(* Logix 5000 project; controller FV vendor 1 type 14 code 217 rev 31.11; software revision 31.00; part 34 of 63 *)
(* tags used below, declared in another part *)
   CheckTimeMask : INT;
   CWD : CHECKWORD_FLAGS;
   Dummy : BOOL;
   FV_A_CTNo : DINT;
   FV_A_CTNo_PLCtoPC : DINT;
   FV_A_FVNo : DINT;
   FV_A_FVNo_PLCtoPC : DINT;
   FV_A_MVNo : DINT;
   FV_A_MVNo_PLCtoPC : DINT;
   FV_ALARM_RETURNED_STRING : STRING;
   FV_Event_Alarm_Tag : ALARM_DIGITAL;
   FV_Event_control_FIFO : CONTROL;
   FV_Event_control_FIFO_Operation_Type : CONTROL;
   FV_Event_Delay_For_Data : TIMER;
   FV_Event_Delay_For_PLC_Startup_Data : TIMER;
   FV_Event_Delay_Timer : TIMER;
   FV_Event_Delay_Timer_Off : TIMER;
   FV_Event_from_buffer : STRING;
   FV_Event_from_buffer_LogData1 : REAL;
   FV_Event_from_buffer_LogData2 : REAL;
   FV_Event_from_buffer_LogData3 : REAL;
   FV_Event_from_buffer_LogData4 : REAL;
   FV_Event_from_buffer_Operation_Type : DINT;
   fv_event_step : DINT;   // 0 - Wait For Event 1 - Sending Event To FactoryTalk 2 - Waiting For Delay Before Next Event Allowed
   FV_Event_String_Last : STRING;
   FV_Event_Transact_Trigger_Tag : DINT;
   FV_Events_FIFO_Buffer : STRING[31];
   FV_Events_FIFO_Buffer_Operation_Type : DINT[31];
   FV_Last_LogData_For_Op : REAL[30,20];
   FV_N20 : INT[255];   // YSVFILL<PC YSV Filling data fro m PC
   FV_N21 : INT[255];   // YSVFILL>PC YSV Filling process data to PC and contr ol regs
   FV_N21_4_alarm : ALARM_DIGITAL;
   FV_N21_4_Alarm_Ready : BOOL;
   FV_N21_4_Delayed_Timer2 : TIMER;
   FV_N21_4_Fault_Returned : STRING;
   FV_N21_4_SQL_Done : DINT;
   FV_N30 : INT[255];   // PITCH<PC YSV Pitching data fr om PC
   FV_N31 : INT[255];   // PITCH>PC YSV Pitching data at o PC and control reg isters
   FV_N31_4_alarm : ALARM_DIGITAL;
   FV_N31_4_Alarm_Ready : BOOL;
   FV_N31_4_Delayed_Timer2 : TIMER;
   FV_N31_4_Fault_Returned : STRING;
   FV_N31_4_SQL_Done : DINT;
   FV_N40 : INT[255];   // YSVCIP<PC
   FV_N41 : INT[255];   // YSVCIP>PC
   FV_N41_4_alarm : ALARM_DIGITAL;
   FV_N41_4_Alarm_Ready : BOOL;
   FV_N41_4_Delayed_Timer2 : TIMER;
   FV_N41_4_Fault_Returned : STRING;
   FV_N41_4_SQL_Done : DINT;
   FV_N50 : INT[255];   // WASTE<PC
   FV_N51 : INT[255];   // WASTE>PC
   FV_N51_4_alarm : ALARM_DIGITAL;
   FV_N51_4_Alarm_Ready : BOOL;
   FV_N51_4_Delayed_Timer2 : TIMER;
   FV_N51_4_Fault_Returned : STRING;
   FV_N51_4_SQL_Done : DINT;
   FV_N60 : INT[255];   // RESEED<PC
   FV_N61 : INT[255];   // RESEED>PC
   FV_N61_4_alarm : ALARM_DIGITAL;
   FV_N61_4_Alarm_Ready : BOOL;
   FV_N61_4_Delayed_Timer2 : TIMER;
   FV_N61_4_Fault_Returned : STRING;
   FV_N61_4_SQL_Done : DINT;
   FV_N71 : INT[255];   // LNCIP >PC
   FV_N71_4_alarm : ALARM_DIGITAL;
   FV_N71_4_Alarm_Ready : BOOL;
   FV_N71_4_Delayed_Timer2 : TIMER;
   FV_N71_4_Fault_Returned : STRING;
   FV_N71_4_SQL_Done : DINT;
   FV_N80 : INT[255];   // YSTFILL<PC YST filling data fro m PC
   FV_N81 : INT[255];   // YSTFILL>PC YST filling process data to PC and contr ol regs.
   FV_N81_4_alarm : ALARM_DIGITAL;
   FV_N81_4_Alarm_Ready : BOOL;
   FV_N81_4_Delayed_Timer2 : TIMER;
   FV_N81_4_Fault_Returned : STRING;
   FV_N81_4_SQL_Done : DINT;
   FV_N84 : INT[255];   // YSTCIP<PC YST CIP data from PC
   FV_N85 : INT[255];   // YSTCIP>PC YST CIP process data to PC and control r egs.
   FV_N85_4_alarm : ALARM_DIGITAL;
   FV_N85_4_Alarm_Ready : BOOL;
   FV_N85_4_Delayed_Timer2 : TIMER;
   FV_N85_4_Fault_Returned : STRING;
   FV_N85_4_SQL_Done : DINT;
   FV_YSTCIP_Log_ID : DINT;
   FV_YSTFILL_Log_ID : DINT;
   FV_YSTs_CIP_Vessel_Event : STRING;
   FV_YSTs_CIP_Vessel_Event_Prefix : STRING;
   FV_YSTs_Filling_Event : STRING;
   FV_YSTs_Filling_Event_Prefix : STRING;
   FV_YSVCIPLINE_Log_ID : DINT;
   FV_YSVCIPVESSEL_Log_ID : DINT;
   FV_YSVFILL_Log_ID : DINT;
   FV_YSVPITCH_Log_ID : DINT;
   FV_YSVRESEED_Log_ID : DINT;
   FV_YSVs_CIP_Line_Event : STRING;
   FV_YSVs_CIP_Line_Event_prefix : STRING;
   FV_YSVs_CIP_vessel_Event : STRING;
   FV_YSVs_CIP_vessel_Event_Prefix : STRING;
   FV_YSVs_Filling_Event : STRING;
   FV_YSVs_Filling_Event_Prefix : STRING;
   FV_YSVs_Pitching_Event : STRING;
   FV_YSVs_Pitching_Event_Prefix : STRING;
   FV_YSVs_reseeding_event : STRING;
   FV_YSVs_reseeding_event_prefix : STRING;
   FV_YSVs_to_waste_event : STRING;
   FV_YSVs_to_waste_event_prefix : STRING;
   FV_YSVTOWASTE_Log_ID : DINT;
(* FV_Common, continued *)

ROUTINE Constants   (* ladder *)
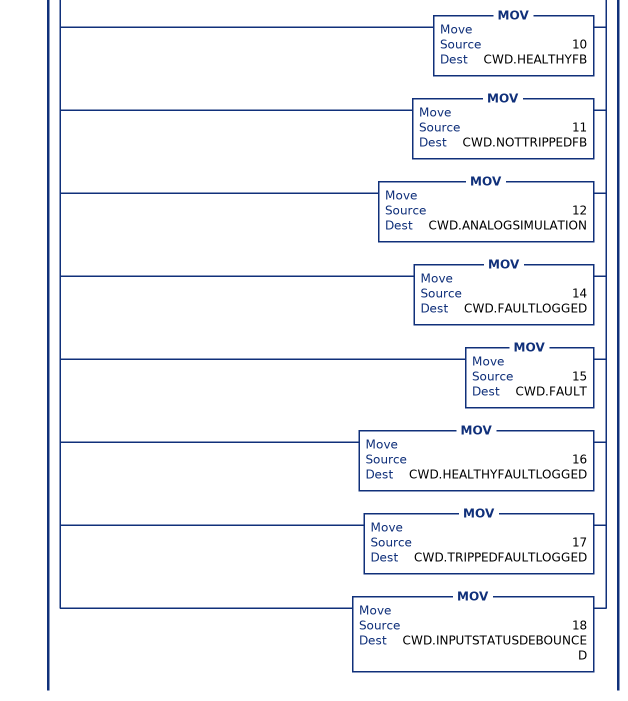
   0: [MOV(0,CWD.AUTODRV) ,MOV(0,CWD.INPUTSTATUS) ,MOV(1,CWD.PREVSCAN) ,MOV(2,CWD.SIMFAIL) ,MOV(3,CWD.OPENFB) ,MOV(3,CWD.RUNFB) ,MOV(4,CWD.CLOSEDFB) ,MOV(5,CWD.MANDRV) ,MOV(6,CWD.MANUAL) ,MOV(7,CWD.OUTPUT) ,MOV(8,CWD.CHECKOFF) ,MOV(9,CWD.HIGHLIGHT) ,MOV(10,CWD.HEALTHYFB) ,MOV(11,CWD.NOTTRIPPEDFB) ,MOV(12,CWD.ANALOGSIMULATION) ,MOV(14,CWD.FAULTLOGGED) ,MOV(15,CWD.FAULT) ,MOV(16,CWD.HEALTHYFAULTLOGGED) ,MOV(17,CWD.TRIPPEDFAULTLOGGED) ,MOV(18,CWD.INPUTSTATUSDEBOUNCED) ];
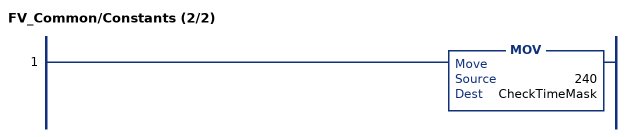
   1: MOV(240,CheckTimeMask);
END_ROUTINE

ROUTINE FV_A_Alarms_From_PLC   (* ladder *)
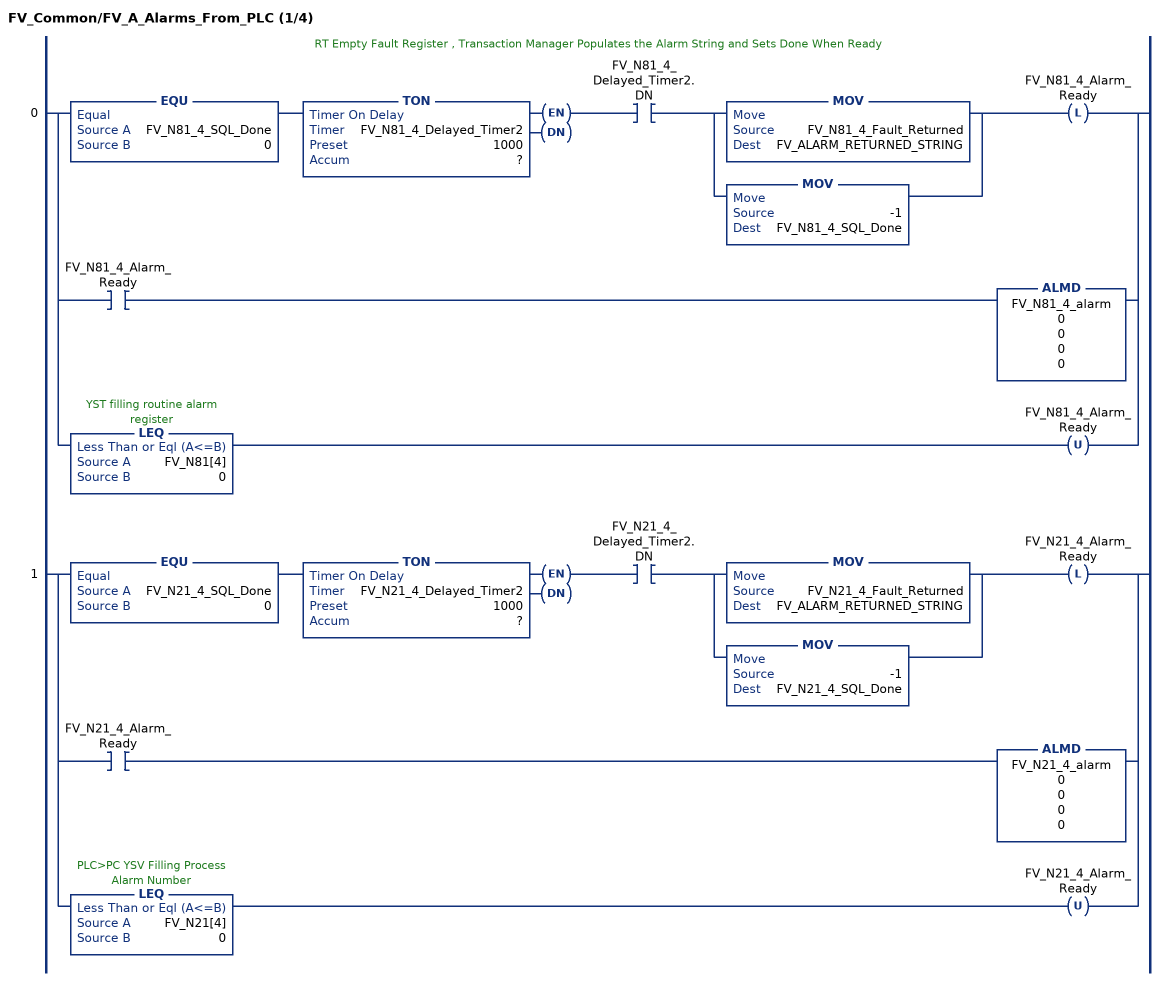
   // RT Empty Fault Register , Transaction Manager Populates the Alarm String and Sets Done When Ready
   0: [EQU(FV_N81_4_SQL_Done,0) TON(FV_N81_4_Delayed_Timer2,?,?) XIC(FV_N81_4_Delayed_Timer2.DN) [MOV(FV_N81_4_Fault_Returned,FV_ALARM_RETURNED_STRING) ,MOV(-1,FV_N81_4_SQL_Done) ] OTL(FV_N81_4_Alarm_Ready) ,XIC(FV_N81_4_Alarm_Ready) ALMD(FV_N81_4_alarm,0,0,0,0) ,LEQ(FV_N81[4],0) OTU(FV_N81_4_Alarm_Ready) ];
   1: [EQU(FV_N21_4_SQL_Done,0) TON(FV_N21_4_Delayed_Timer2,?,?) XIC(FV_N21_4_Delayed_Timer2.DN) [MOV(FV_N21_4_Fault_Returned,FV_ALARM_RETURNED_STRING) ,MOV(-1,FV_N21_4_SQL_Done) ] OTL(FV_N21_4_Alarm_Ready) ,XIC(FV_N21_4_Alarm_Ready) ALMD(FV_N21_4_alarm,0,0,0,0) ,LEQ(FV_N21[4],0) OTU(FV_N21_4_Alarm_Ready) ];
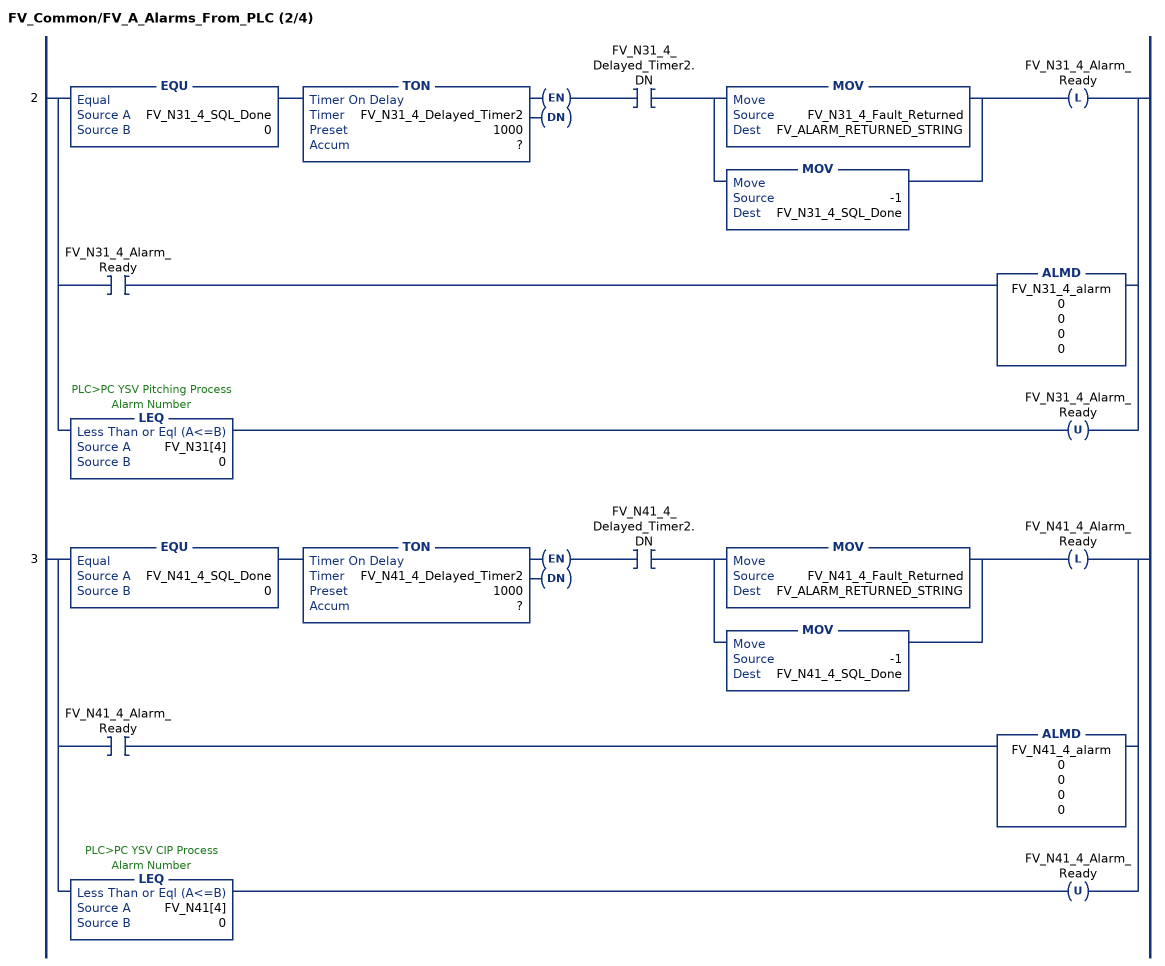
   2: [EQU(FV_N31_4_SQL_Done,0) TON(FV_N31_4_Delayed_Timer2,?,?) XIC(FV_N31_4_Delayed_Timer2.DN) [MOV(FV_N31_4_Fault_Returned,FV_ALARM_RETURNED_STRING) ,MOV(-1,FV_N31_4_SQL_Done) ] OTL(FV_N31_4_Alarm_Ready) ,XIC(FV_N31_4_Alarm_Ready) ALMD(FV_N31_4_alarm,0,0,0,0) ,LEQ(FV_N31[4],0) OTU(FV_N31_4_Alarm_Ready) ];
   3: [EQU(FV_N41_4_SQL_Done,0) TON(FV_N41_4_Delayed_Timer2,?,?) XIC(FV_N41_4_Delayed_Timer2.DN) [MOV(FV_N41_4_Fault_Returned,FV_ALARM_RETURNED_STRING) ,MOV(-1,FV_N41_4_SQL_Done) ] OTL(FV_N41_4_Alarm_Ready) ,XIC(FV_N41_4_Alarm_Ready) ALMD(FV_N41_4_alarm,0,0,0,0) ,LEQ(FV_N41[4],0) OTU(FV_N41_4_Alarm_Ready) ];
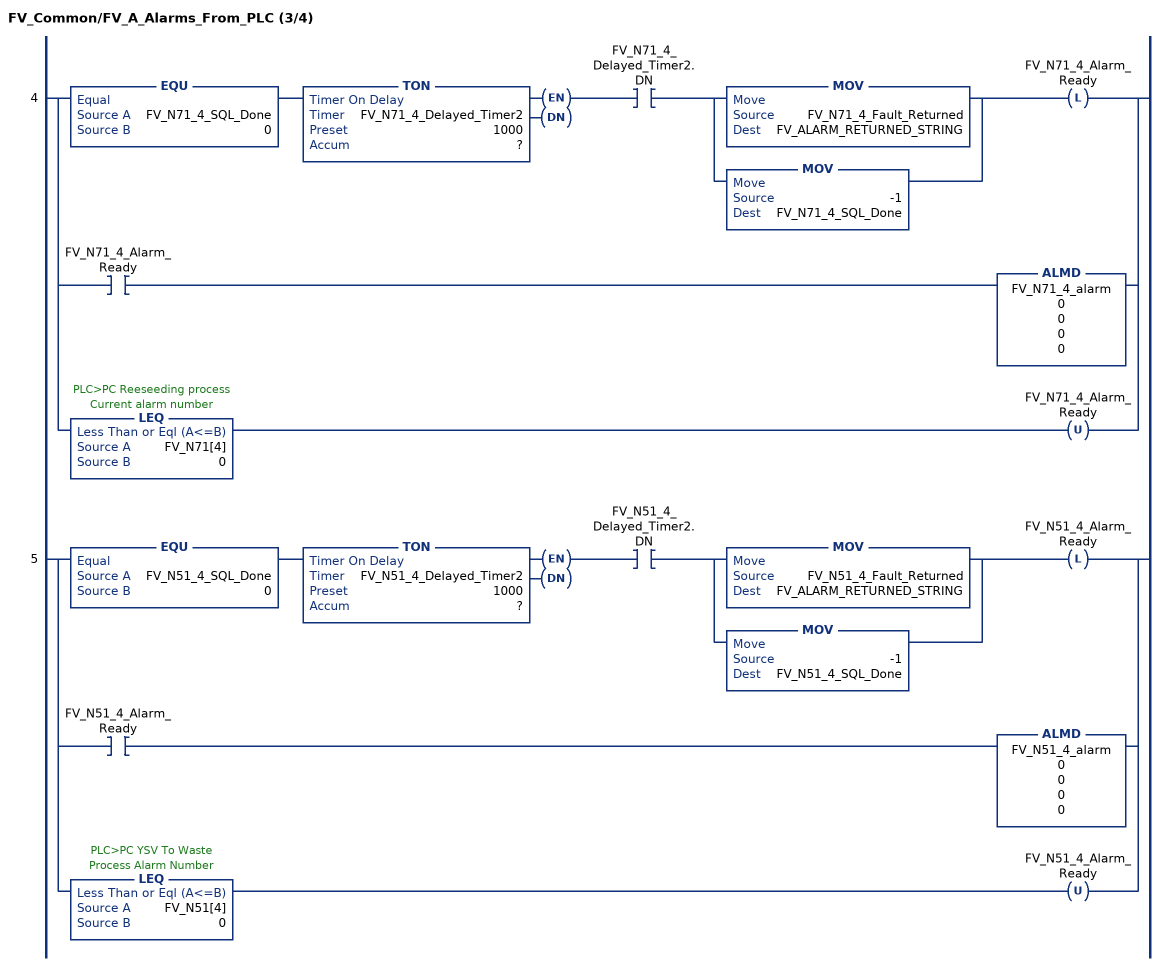
   4: [EQU(FV_N71_4_SQL_Done,0) TON(FV_N71_4_Delayed_Timer2,?,?) XIC(FV_N71_4_Delayed_Timer2.DN) [MOV(FV_N71_4_Fault_Returned,FV_ALARM_RETURNED_STRING) ,MOV(-1,FV_N71_4_SQL_Done) ] OTL(FV_N71_4_Alarm_Ready) ,XIC(FV_N71_4_Alarm_Ready) ALMD(FV_N71_4_alarm,0,0,0,0) ,LEQ(FV_N71[4],0) OTU(FV_N71_4_Alarm_Ready) ];
   5: [EQU(FV_N51_4_SQL_Done,0) TON(FV_N51_4_Delayed_Timer2,?,?) XIC(FV_N51_4_Delayed_Timer2.DN) [MOV(FV_N51_4_Fault_Returned,FV_ALARM_RETURNED_STRING) ,MOV(-1,FV_N51_4_SQL_Done) ] OTL(FV_N51_4_Alarm_Ready) ,XIC(FV_N51_4_Alarm_Ready) ALMD(FV_N51_4_alarm,0,0,0,0) ,LEQ(FV_N51[4],0) OTU(FV_N51_4_Alarm_Ready) ];
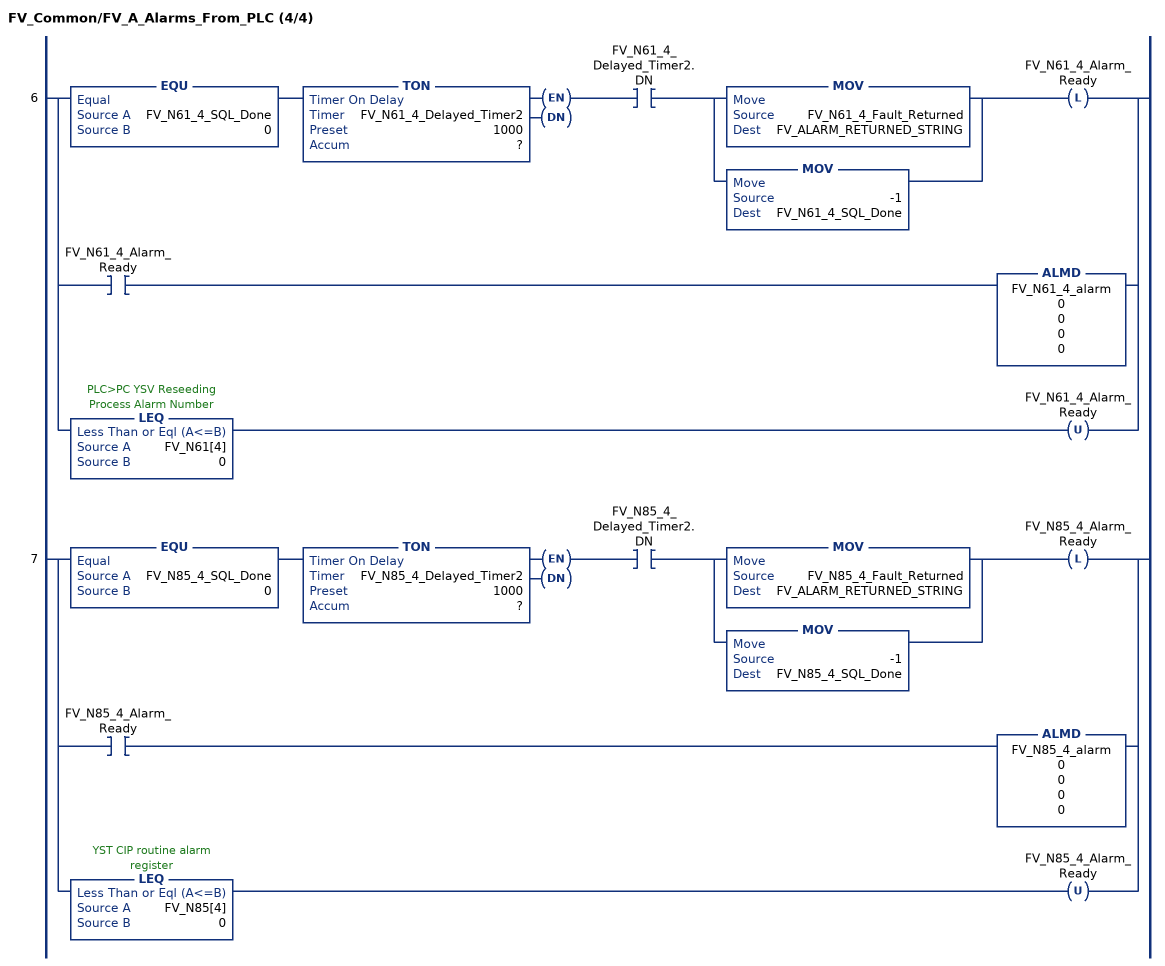
   6: [EQU(FV_N61_4_SQL_Done,0) TON(FV_N61_4_Delayed_Timer2,?,?) XIC(FV_N61_4_Delayed_Timer2.DN) [MOV(FV_N61_4_Fault_Returned,FV_ALARM_RETURNED_STRING) ,MOV(-1,FV_N61_4_SQL_Done) ] OTL(FV_N61_4_Alarm_Ready) ,XIC(FV_N61_4_Alarm_Ready) ALMD(FV_N61_4_alarm,0,0,0,0) ,LEQ(FV_N61[4],0) OTU(FV_N61_4_Alarm_Ready) ];
   7: [EQU(FV_N85_4_SQL_Done,0) TON(FV_N85_4_Delayed_Timer2,?,?) XIC(FV_N85_4_Delayed_Timer2.DN) [MOV(FV_N85_4_Fault_Returned,FV_ALARM_RETURNED_STRING) ,MOV(-1,FV_N85_4_SQL_Done) ] OTL(FV_N85_4_Alarm_Ready) ,XIC(FV_N85_4_Alarm_Ready) ALMD(FV_N85_4_alarm,0,0,0,0) ,LEQ(FV_N85[4],0) OTU(FV_N85_4_Alarm_Ready) ];
END_ROUTINE

ROUTINE FV_A_CTNo_PLCtoPC   (* ladder *)
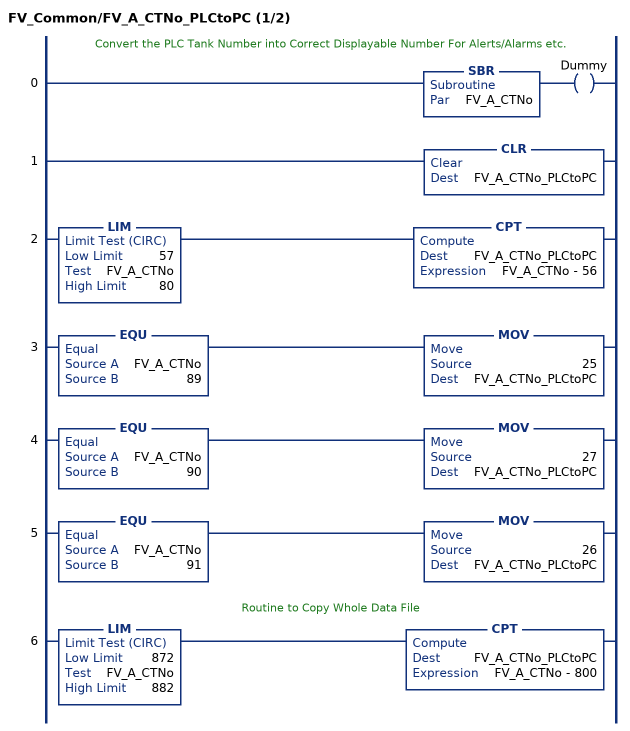
   // Convert the PLC Tank Number into Correct Displayable Number For Alerts/Alarms etc.
   0: SBR(FV_A_CTNo)OTE(Dummy);
   1: CLR(FV_A_CTNo_PLCtoPC);
   2: LIM(57,FV_A_CTNo,80)CPT(FV_A_CTNo_PLCtoPC,FV_A_CTNo - 56);
   3: EQU(FV_A_CTNo,89)MOV(25,FV_A_CTNo_PLCtoPC);
   4: EQU(FV_A_CTNo,90)MOV(27,FV_A_CTNo_PLCtoPC);
   5: EQU(FV_A_CTNo,91)MOV(26,FV_A_CTNo_PLCtoPC);
   // Routine to Copy Whole Data File
   6: LIM(872,FV_A_CTNo,882)CPT(FV_A_CTNo_PLCtoPC,FV_A_CTNo - 800);
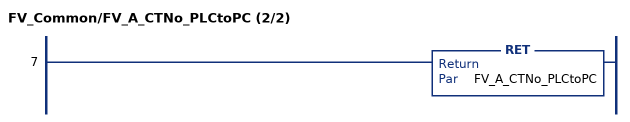
   7: RET(FV_A_CTNo_PLCtoPC);
END_ROUTINE

ROUTINE FV_A_Events_From_Scada   (* ladder *)
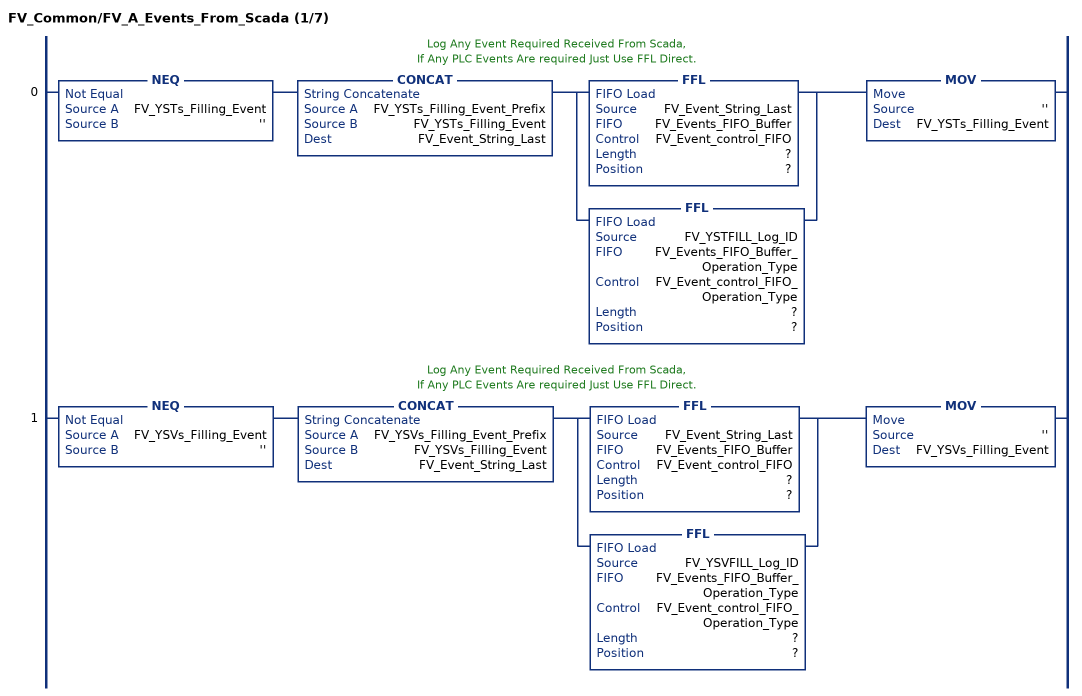
   // Log Any Event Required Received From Scada,
   // If Any PLC Events Are required Just Use FFL Direct.
   0: NEQ(FV_YSTs_Filling_Event,'')CONCAT(FV_YSTs_Filling_Event_Prefix,FV_YSTs_Filling_Event,FV_Event_String_Last)[FFL(FV_Event_String_Last,FV_Events_FIFO_Buffer,FV_Event_control_FIFO,?,?) ,FFL(FV_YSTFILL_Log_ID,FV_Events_FIFO_Buffer_Operation_Type,FV_Event_control_FIFO_Operation_Type,?,?) ]MOV('',FV_YSTs_Filling_Event);
   // Log Any Event Required Received From Scada,
   // If Any PLC Events Are required Just Use FFL Direct.
   1: NEQ(FV_YSVs_Filling_Event,'')CONCAT(FV_YSVs_Filling_Event_Prefix,FV_YSVs_Filling_Event,FV_Event_String_Last)[FFL(FV_Event_String_Last,FV_Events_FIFO_Buffer,FV_Event_control_FIFO,?,?) ,FFL(FV_YSVFILL_Log_ID,FV_Events_FIFO_Buffer_Operation_Type,FV_Event_control_FIFO_Operation_Type,?,?) ]MOV('',FV_YSVs_Filling_Event);
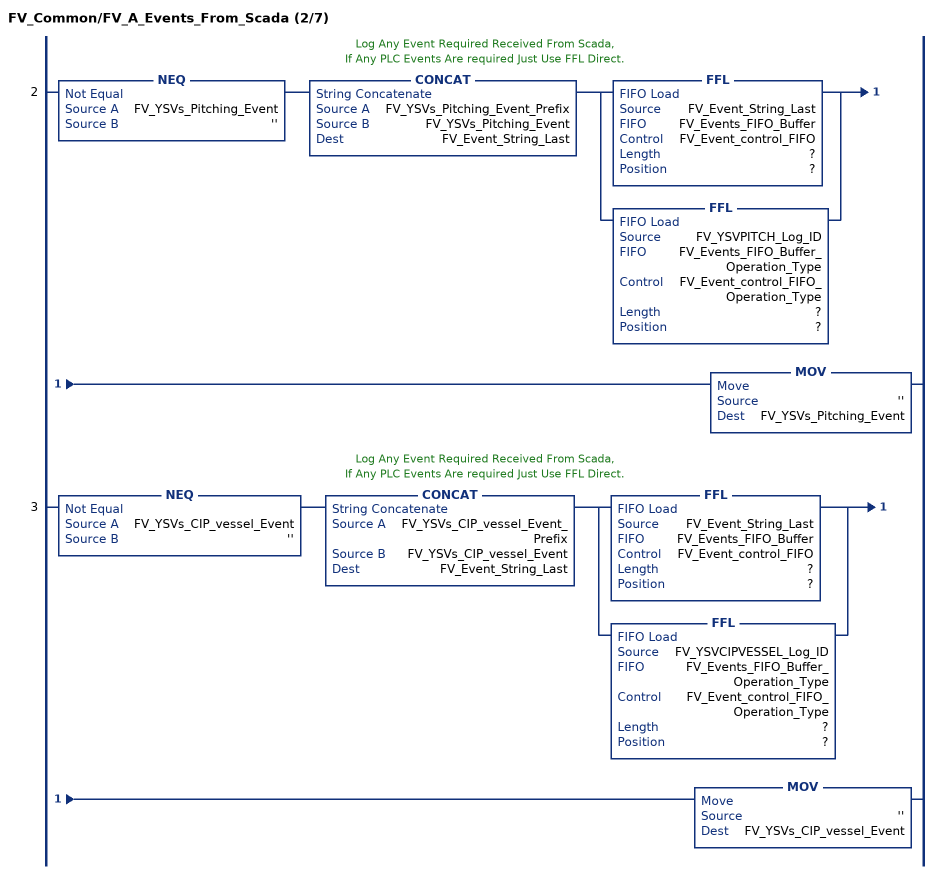
   // Log Any Event Required Received From Scada,
   // If Any PLC Events Are required Just Use FFL Direct.
   2: NEQ(FV_YSVs_Pitching_Event,'')CONCAT(FV_YSVs_Pitching_Event_Prefix,FV_YSVs_Pitching_Event,FV_Event_String_Last)[FFL(FV_Event_String_Last,FV_Events_FIFO_Buffer,FV_Event_control_FIFO,?,?) ,FFL(FV_YSVPITCH_Log_ID,FV_Events_FIFO_Buffer_Operation_Type,FV_Event_control_FIFO_Operation_Type,?,?) ]MOV('',FV_YSVs_Pitching_Event);
   // Log Any Event Required Received From Scada,
   // If Any PLC Events Are required Just Use FFL Direct.
   3: NEQ(FV_YSVs_CIP_vessel_Event,'')CONCAT(FV_YSVs_CIP_vessel_Event_Prefix,FV_YSVs_CIP_vessel_Event,FV_Event_String_Last)[FFL(FV_Event_String_Last,FV_Events_FIFO_Buffer,FV_Event_control_FIFO,?,?) ,FFL(FV_YSVCIPVESSEL_Log_ID,FV_Events_FIFO_Buffer_Operation_Type,FV_Event_control_FIFO_Operation_Type,?,?) ]MOV('',FV_YSVs_CIP_vessel_Event);
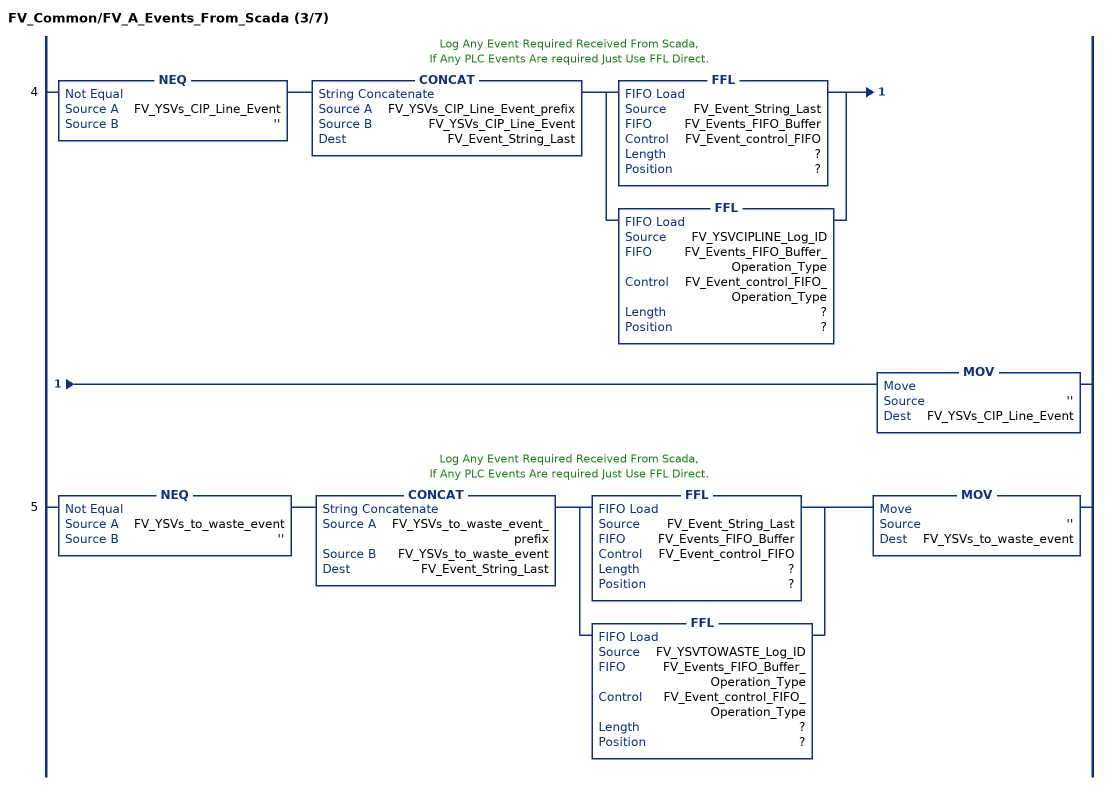
   // Log Any Event Required Received From Scada,
   // If Any PLC Events Are required Just Use FFL Direct.
   4: NEQ(FV_YSVs_CIP_Line_Event,'')CONCAT(FV_YSVs_CIP_Line_Event_prefix,FV_YSVs_CIP_Line_Event,FV_Event_String_Last)[FFL(FV_Event_String_Last,FV_Events_FIFO_Buffer,FV_Event_control_FIFO,?,?) ,FFL(FV_YSVCIPLINE_Log_ID,FV_Events_FIFO_Buffer_Operation_Type,FV_Event_control_FIFO_Operation_Type,?,?) ]MOV('',FV_YSVs_CIP_Line_Event);
   // Log Any Event Required Received From Scada,
   // If Any PLC Events Are required Just Use FFL Direct.
   5: NEQ(FV_YSVs_to_waste_event,'')CONCAT(FV_YSVs_to_waste_event_prefix,FV_YSVs_to_waste_event,FV_Event_String_Last)[FFL(FV_Event_String_Last,FV_Events_FIFO_Buffer,FV_Event_control_FIFO,?,?) ,FFL(FV_YSVTOWASTE_Log_ID,FV_Events_FIFO_Buffer_Operation_Type,FV_Event_control_FIFO_Operation_Type,?,?) ]MOV('',FV_YSVs_to_waste_event);
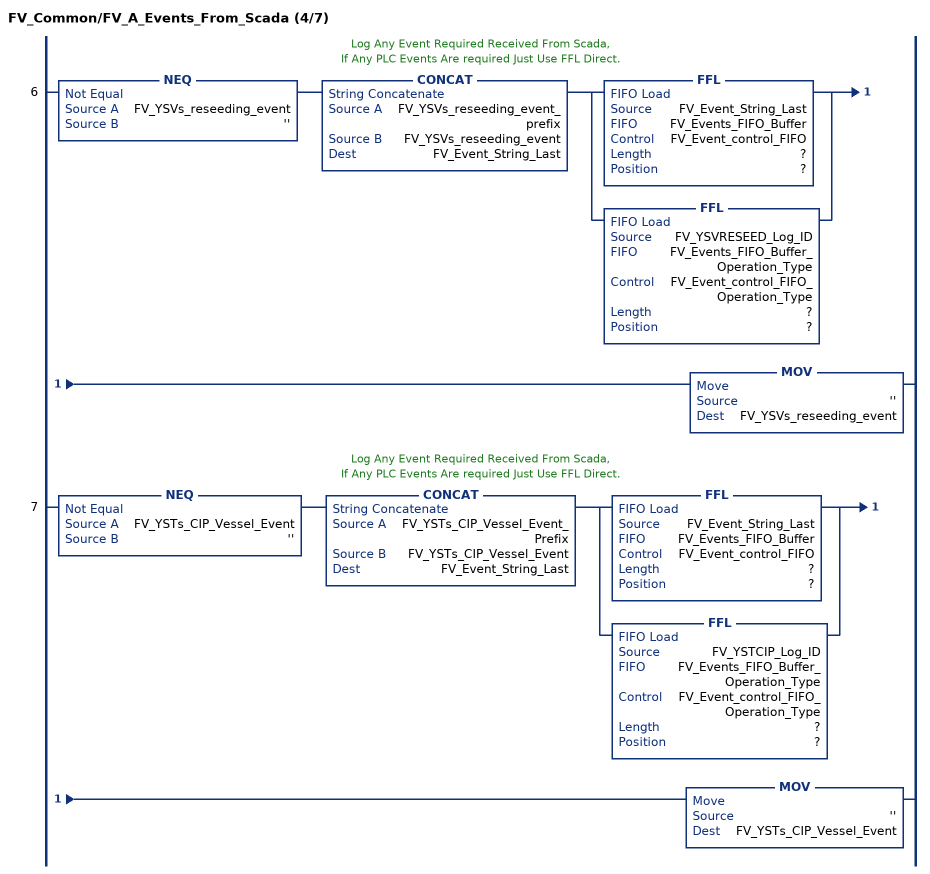
   // Log Any Event Required Received From Scada,
   // If Any PLC Events Are required Just Use FFL Direct.
   6: NEQ(FV_YSVs_reseeding_event,'')CONCAT(FV_YSVs_reseeding_event_prefix,FV_YSVs_reseeding_event,FV_Event_String_Last)[FFL(FV_Event_String_Last,FV_Events_FIFO_Buffer,FV_Event_control_FIFO,?,?) ,FFL(FV_YSVRESEED_Log_ID,FV_Events_FIFO_Buffer_Operation_Type,FV_Event_control_FIFO_Operation_Type,?,?) ]MOV('',FV_YSVs_reseeding_event);
   // Log Any Event Required Received From Scada,
   // If Any PLC Events Are required Just Use FFL Direct.
   7: NEQ(FV_YSTs_CIP_Vessel_Event,'')CONCAT(FV_YSTs_CIP_Vessel_Event_Prefix,FV_YSTs_CIP_Vessel_Event,FV_Event_String_Last)[FFL(FV_Event_String_Last,FV_Events_FIFO_Buffer,FV_Event_control_FIFO,?,?) ,FFL(FV_YSTCIP_Log_ID,FV_Events_FIFO_Buffer_Operation_Type,FV_Event_control_FIFO_Operation_Type,?,?) ]MOV('',FV_YSTs_CIP_Vessel_Event);
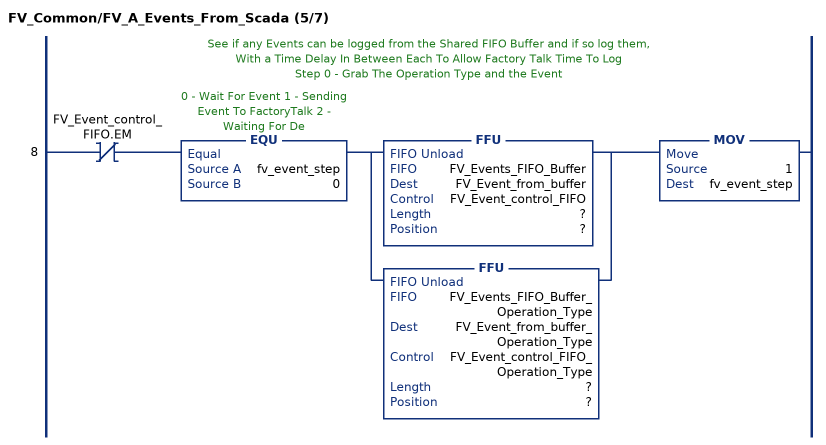
   // See if any Events can be logged from the Shared FIFO Buffer and if so log them,
   // With a Time Delay In Between Each To Allow Factory Talk Time To Log
   // Step 0 - Grab The Operation Type and the Event
   8: XIO(FV_Event_control_FIFO.EM)EQU(fv_event_step,0)[FFU(FV_Events_FIFO_Buffer,FV_Event_from_buffer,FV_Event_control_FIFO,?,?) ,FFU(FV_Events_FIFO_Buffer_Operation_Type,FV_Event_from_buffer_Operation_Type,FV_Event_control_FIFO_Operation_Type,?,?) ]MOV(1,fv_event_step);
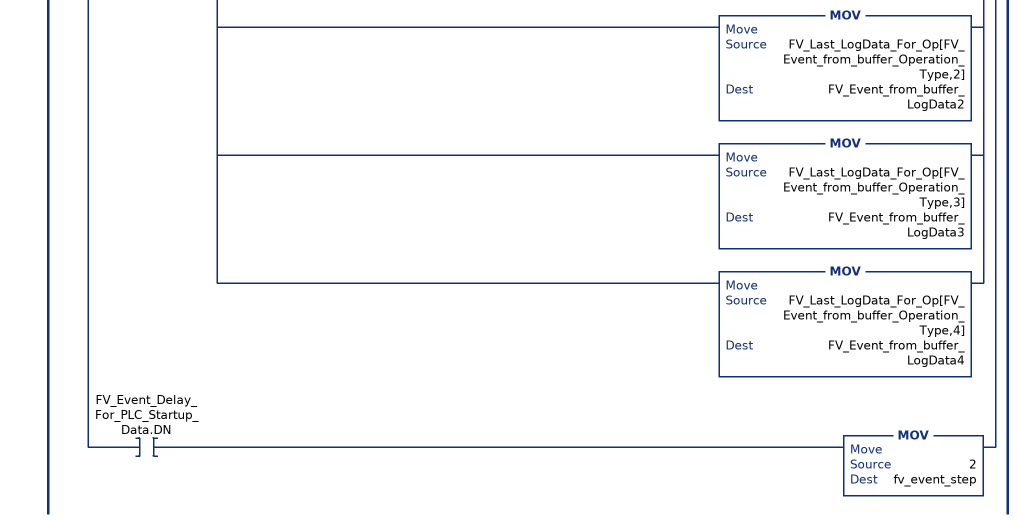
   // Wait For PLC To Shift The Data, Especially important on Startup as the Start event is from the PC and the Data is only put in place when the PLC Starts the operation.
   // Also Stores Last If Required, As Abort will have the data wiped out prior to event being logged
   9: EQU(fv_event_step,1)[TON(FV_Event_Delay_For_PLC_Startup_Data,?,?) ,CLR(FV_Event_from_buffer_LogData1) CLR(FV_Event_from_buffer_LogData2) CLR(FV_Event_from_buffer_LogData3) CLR(FV_Event_from_buffer_LogData4) ,XIC(FV_Event_Delay_For_PLC_Startup_Data.DN) [EQU(FV_Event_from_buffer_Operation_Type,FV_YSTFILL_Log_ID) GRT(FV_N80[1],0) ADD(FV_N80[1],94,FV_Last_LogData_For_Op[FV_Event_from_buffer_Operation_Type,2]) ,EQU(FV_Event_from_buffer_Operation_Type,FV_YSVFILL_Log_ID) GRT(FV_N20[1],0) ADD(FV_N20[1],25,FV_Last_LogData_For_Op[FV_Event_from_buffer_Operation_Type,2]) ,EQU(FV_Event_from_buffer_Operation_Type,FV_YSVPITCH_Log_ID) [GRT(FV_N30[1],0) ADD(FV_N30[1],25,FV_Last_LogData_For_Op[FV_Event_from_buffer_Operation_Type,1]) ,GRT(FV_N30[3],0) MOV(FV_N30[3],FV_Last_LogData_For_Op[FV_Event_from_buffer_Operation_Type,2]) ] ,EQU(FV_Event_from_buffer_Operation_Type,FV_YSVCIPVESSEL_Log_ID) GRT(FV_N40[1],0) ADD(FV_N40[1],25,FV_Last_LogData_For_Op[FV_Event_from_buffer_Operation_Type,1]) ,EQU(FV_Event_from_buffer_Operation_Type,FV_YSVCIPLINE_Log_ID) MOV(0,FV_Last_LogData_For_Op[FV_Event_from_buffer_Operation_Type,1]) ,EQU(FV_Event_from_buffer_Operation_Type,FV_YSVTOWASTE_Log_ID) GRT(FV_N50[1],0) ADD(FV_N50[1],25,FV_Last_LogData_For_Op[FV_Event_from_buffer_Operation_Type,1]) ,EQU(FV_Event_from_buffer_Operation_Type,FV_YSVRESEED_Log_ID) [GRT(FV_N60[3],0) MOV(FV_N60[3],FV_Last_LogData_For_Op[FV_Event_from_buffer_Operation_Type,1]) ,GRT(FV_N60[4],0) MOV(FV_N60[4],FV_Last_LogData_For_Op[FV_Event_from_buffer_Operation_Type,2]) ] ,EQU(FV_Event_from_buffer_Operation_Type,FV_YSTCIP_Log_ID) GRT(FV_N84[1],0) ADD(FV_N84[1],94,FV_Last_LogData_For_Op[FV_Event_from_buffer_Operation_Type,1]) ] ,XIC(FV_Event_Delay_For_PLC_Startup_Data.DN) [MOV(FV_Last_LogData_For_Op[FV_Event_from_buffer_Operation_Type,1],FV_Event_from_buffer_LogData1) ,MOV(FV_Last_LogData_For_Op[FV_Event_from_buffer_Operation_Type,2],FV_Event_from_buffer_LogData2) ,MOV(FV_Last_LogData_For_Op[FV_Event_from_buffer_Operation_Type,3],FV_Event_from_buffer_LogData3) ,MOV(FV_Last_LogData_For_Op[FV_Event_from_buffer_Operation_Type,4],FV_Event_from_buffer_LogData4) ] ,XIC(FV_Event_Delay_For_PLC_Startup_Data.DN) MOV(2,fv_event_step) ];
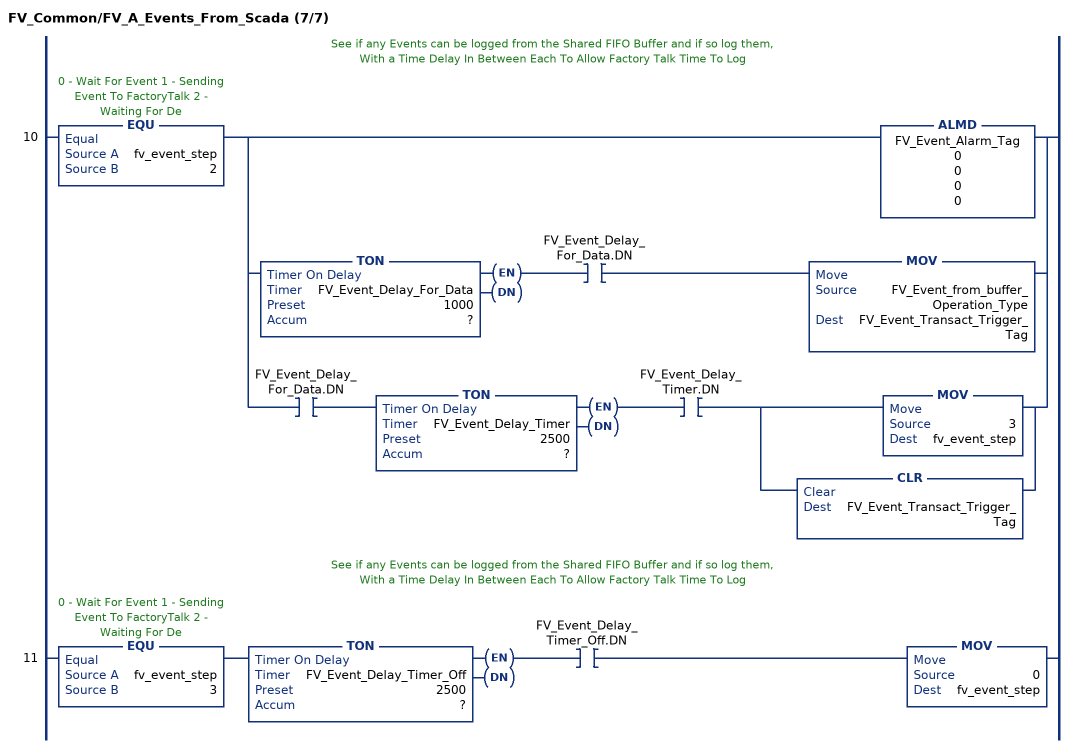
   // See if any Events can be logged from the Shared FIFO Buffer and if so log them,
   // With a Time Delay In Between Each To Allow Factory Talk Time To Log
   10: EQU(fv_event_step,2)[ALMD(FV_Event_Alarm_Tag,0,0,0,0) ,TON(FV_Event_Delay_For_Data,?,?) XIC(FV_Event_Delay_For_Data.DN) MOV(FV_Event_from_buffer_Operation_Type,FV_Event_Transact_Trigger_Tag) ,XIC(FV_Event_Delay_For_Data.DN) TON(FV_Event_Delay_Timer,?,?) XIC(FV_Event_Delay_Timer.DN) [MOV(3,fv_event_step) ,CLR(FV_Event_Transact_Trigger_Tag) ] ];
   // See if any Events can be logged from the Shared FIFO Buffer and if so log them,
   // With a Time Delay In Between Each To Allow Factory Talk Time To Log
   11: EQU(fv_event_step,3)TON(FV_Event_Delay_Timer_Off,?,?)XIC(FV_Event_Delay_Timer_Off.DN)MOV(0,fv_event_step);
END_ROUTINE

ROUTINE FV_A_Events_From_Scada_IDs   (* ladder *)
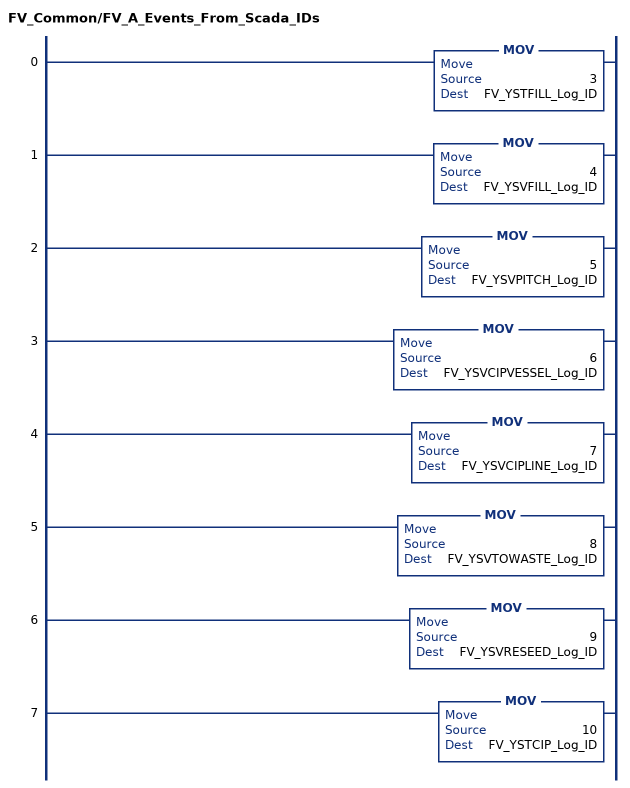
   0: MOV(3,FV_YSTFILL_Log_ID);
   1: MOV(4,FV_YSVFILL_Log_ID);
   2: MOV(5,FV_YSVPITCH_Log_ID);
   3: MOV(6,FV_YSVCIPVESSEL_Log_ID);
   4: MOV(7,FV_YSVCIPLINE_Log_ID);
   5: MOV(8,FV_YSVTOWASTE_Log_ID);
   6: MOV(9,FV_YSVRESEED_Log_ID);
   7: MOV(10,FV_YSTCIP_Log_ID);
END_ROUTINE

ROUTINE FV_A_FVNo_PLCtoPC   (* ladder *)
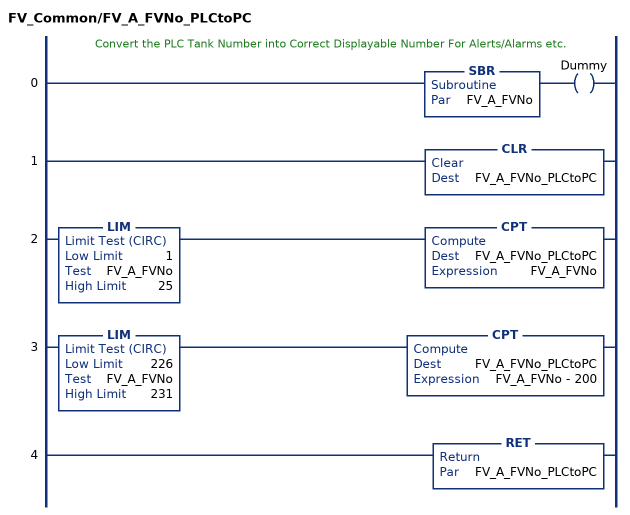
   // Convert the PLC Tank Number into Correct Displayable Number For Alerts/Alarms etc.
   0: SBR(FV_A_FVNo)OTE(Dummy);
   1: CLR(FV_A_FVNo_PLCtoPC);
   2: LIM(1,FV_A_FVNo,25)CPT(FV_A_FVNo_PLCtoPC,FV_A_FVNo);
   3: LIM(226,FV_A_FVNo,231)CPT(FV_A_FVNo_PLCtoPC,FV_A_FVNo - 200);
   4: RET(FV_A_FVNo_PLCtoPC);
END_ROUTINE

ROUTINE FV_A_MVNo_PLCtoPC   (* ladder *)
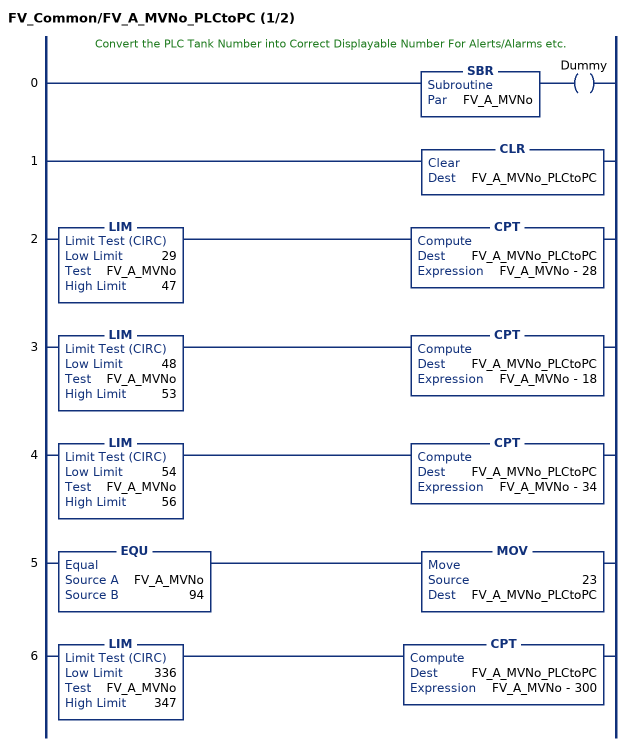
   // Convert the PLC Tank Number into Correct Displayable Number For Alerts/Alarms etc.
   0: SBR(FV_A_MVNo)OTE(Dummy);
   1: CLR(FV_A_MVNo_PLCtoPC);
   2: LIM(29,FV_A_MVNo,47)CPT(FV_A_MVNo_PLCtoPC,FV_A_MVNo - 28);
   3: LIM(48,FV_A_MVNo,53)CPT(FV_A_MVNo_PLCtoPC,FV_A_MVNo - 18);
   4: LIM(54,FV_A_MVNo,56)CPT(FV_A_MVNo_PLCtoPC,FV_A_MVNo - 34);
   5: EQU(FV_A_MVNo,94)MOV(23,FV_A_MVNo_PLCtoPC);
   6: LIM(336,FV_A_MVNo,347)CPT(FV_A_MVNo_PLCtoPC,FV_A_MVNo - 300);
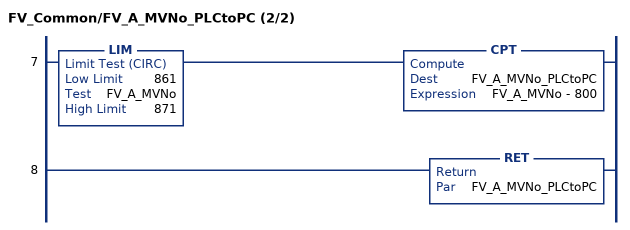
   7: LIM(861,FV_A_MVNo,871)CPT(FV_A_MVNo_PLCtoPC,FV_A_MVNo - 800);
   8: RET(FV_A_MVNo_PLCtoPC);
END_ROUTINE
